// TIA Portal project "GzyHzy_1500" (V15) (continued)
VERSION : 0.1
   VAR
      "1#除尘轴伸端U1相" : Real;   // 临时占位符变量
      "1#除尘轴伸端V1相" : Real;   // 临时占位符变量
      "1#除尘轴伸端W1相" : Real;   // 临时占位符变量
      "1#除尘非轴伸端U2相" : Real;   // 临时占位符变量
      "1#除尘非轴伸端V2相" : Real;   // 临时占位符变量
      "1#除尘非轴伸端W2相" : Real;   // 临时占位符变量
      "1#除尘电机前轴承温度" : Real;   // 临时占位符变量
      "1#除尘电机后轴承温度" : Real;   // 临时占位符变量
      "1#除尘风机前轴承温度" : Real;   // 临时占位符变量
      "1#除尘风机后轴承温度" : Real;   // 临时占位符变量
      DB_VAR10 : Real;   // 临时占位符变量
      DB_VAR11 : Real;   // 临时占位符变量
      DB_VAR12 : Real;   // 临时占位符变量
      DB_VAR13 : Real;   // 临时占位符变量
      DB_VAR14 : Real;   // 临时占位符变量
      DB_VAR15 : Real;   // 临时占位符变量
      DB_VAR16 : Real;   // 临时占位符变量
      DB_VAR17 : Real;   // 临时占位符变量
      DB_VAR18 : Real;   // 临时占位符变量
      DB_VAR19 : Real;   // 临时占位符变量
      DB_VAR20 : Real;   // 临时占位符变量
      DB_VAR21 : Real;   // 临时占位符变量
      DB_VAR22 : Real;   // 临时占位符变量
      DB_VAR23 : Real;   // 临时占位符变量
      DB_VAR24 : Real;   // 临时占位符变量
      DB_VAR25 : Real;   // 临时占位符变量
      DB_VAR26 : Real;   // 临时占位符变量
      DB_VAR27 : Real;   // 临时占位符变量
      DB_VAR28 : Real;   // 临时占位符变量
      DB_VAR29 : Real;   // 临时占位符变量
      DB_VAR30 : Real;   // 临时占位符变量
      DB_VAR31 : Real;   // 临时占位符变量
      DB_VAR32 : Real;   // 临时占位符变量
      DB_VAR33 : Real;   // 临时占位符变量
      DB_VAR34 : Real;   // 临时占位符变量
      DB_VAR35 : Real;   // 临时占位符变量
      DB_VAR36 : Real;   // 临时占位符变量
      DB_VAR37 : Real;   // 临时占位符变量
      DB_VAR38 : Real;   // 临时占位符变量
      DB_VAR39 : Real;   // 临时占位符变量
      DB_VAR40 : Real;   // 临时占位符变量
      DB_VAR41 : Real;   // 临时占位符变量
      DB_VAR42 : Real;   // 临时占位符变量
      DB_VAR43 : Real;   // 临时占位符变量
      DB_VAR44 : Real;   // 临时占位符变量
      DB_VAR45 : Real;   // 临时占位符变量
      DB_VAR46 : Real;   // 临时占位符变量
      DB_VAR47 : Real;   // 临时占位符变量
      DB_VAR48 : Real;   // 临时占位符变量
      DB_VAR49 : Real;   // 临时占位符变量
      "2#除尘轴伸端U1相" : Real;   // 临时占位符变量
      "2#除尘轴伸端V1相" : Real;   // 临时占位符变量
      "2#除尘轴伸端W1相" : Real;   // 临时占位符变量
      "2#除尘非轴伸端U2相" : Real;   // 临时占位符变量
      "2#除尘非轴伸端V2相" : Real;   // 临时占位符变量
      "2#除尘非轴伸端W2相" : Real;   // 临时占位符变量
      "2#除尘电机前轴承温度" : Real;   // 临时占位符变量
      "2#除尘电机后轴承温度" : Real;   // 临时占位符变量
      "2#除尘风机前轴承温度" : Real;   // 临时占位符变量
      "2#除尘风机后轴承温度" : Real;   // 临时占位符变量
      DB_VAR60 : Real;   // 临时占位符变量
      DB_VAR61 : Real;   // 临时占位符变量
      DB_VAR62 : Real;   // 临时占位符变量
      DB_VAR63 : Real;   // 临时占位符变量
      DB_VAR64 : Real;   // 临时占位符变量
      DB_VAR65 : Real;   // 临时占位符变量
      DB_VAR66 : Real;   // 临时占位符变量
   END_VAR
BEGIN
END_DATA_BLOCK

FUNCTION "FC1" : Void   // FC1, LAD
{ S7_Optimized_Access := 'FALSE' }
VERSION : 0.1
BEGIN

REGION Network 1: 1#1号电场二次运行电压
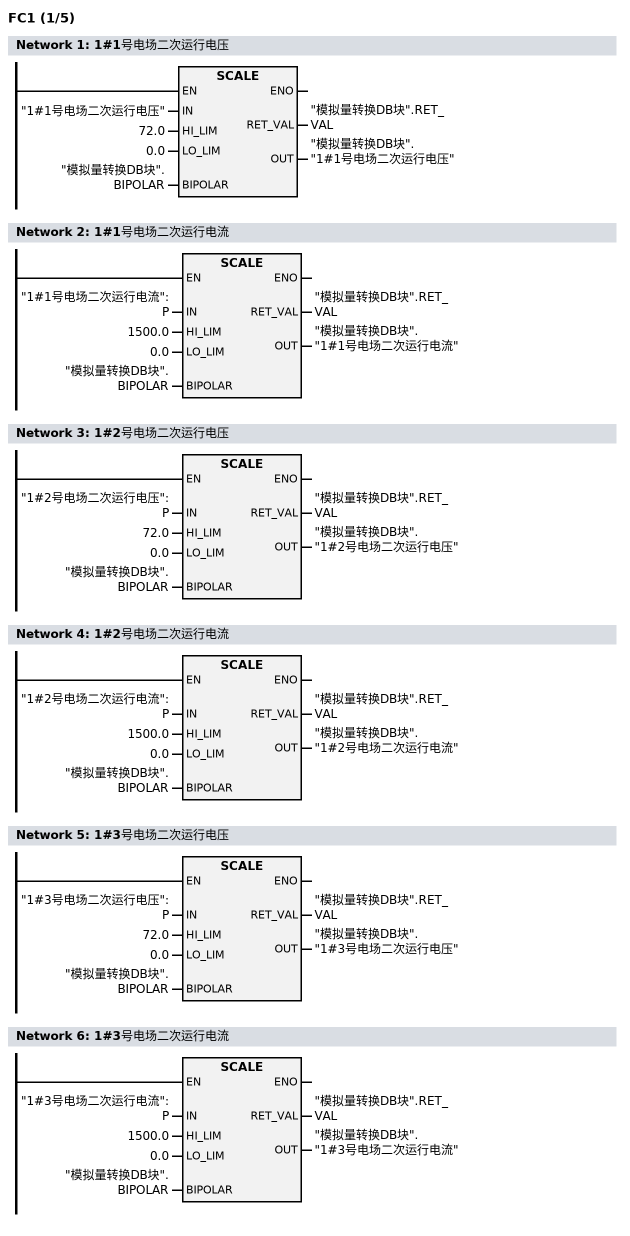
   "模拟量转换DB块".RET_VAL := SCALE(IN := "1#1号电场二次运行电压",
                           HI_LIM := 72.0,
                           LO_LIM := 0.0,
                           BIPOLAR := "模拟量转换DB块".BIPOLAR,
                           OUT => "模拟量转换DB块"."1#1号电场二次运行电压");
END_REGION

REGION Network 2: 1#1号电场二次运行电流
   "模拟量转换DB块".RET_VAL := SCALE(IN := "1#1号电场二次运行电流":P,
                           HI_LIM := 1500.0,
                           LO_LIM := 0.0,
                           BIPOLAR := "模拟量转换DB块".BIPOLAR,
                           OUT => "模拟量转换DB块"."1#1号电场二次运行电流");
END_REGION

REGION Network 3: 1#2号电场二次运行电压
   "模拟量转换DB块".RET_VAL := SCALE(IN := "1#2号电场二次运行电压":P,
                           HI_LIM := 72.0,
                           LO_LIM := 0.0,
                           BIPOLAR := "模拟量转换DB块".BIPOLAR,
                           OUT => "模拟量转换DB块"."1#2号电场二次运行电压");
END_REGION

REGION Network 4: 1#2号电场二次运行电流
   "模拟量转换DB块".RET_VAL := SCALE(IN := "1#2号电场二次运行电流":P,
                           HI_LIM := 1500.0,
                           LO_LIM := 0.0,
                           BIPOLAR := "模拟量转换DB块".BIPOLAR,
                           OUT => "模拟量转换DB块"."1#2号电场二次运行电流");
END_REGION

REGION Network 5: 1#3号电场二次运行电压
   "模拟量转换DB块".RET_VAL := SCALE(IN := "1#3号电场二次运行电压":P,
                           HI_LIM := 72.0,
                           LO_LIM := 0.0,
                           BIPOLAR := "模拟量转换DB块".BIPOLAR,
                           OUT => "模拟量转换DB块"."1#3号电场二次运行电压");
END_REGION

REGION Network 6: 1#3号电场二次运行电流
   "模拟量转换DB块".RET_VAL := SCALE(IN := "1#3号电场二次运行电流":P,
                           HI_LIM := 1500.0,
                           LO_LIM := 0.0,
                           BIPOLAR := "模拟量转换DB块".BIPOLAR,
                           OUT => "模拟量转换DB块"."1#3号电场二次运行电流");
END_REGION

REGION Network 7: 1#4号电场二次运行电压
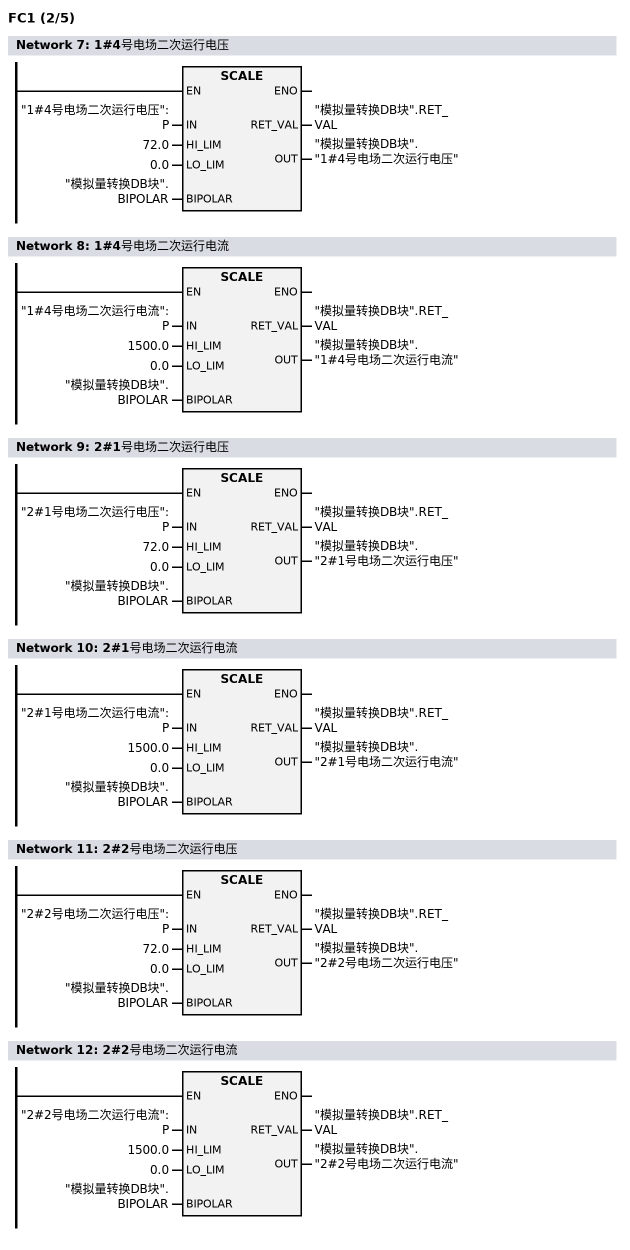
   "模拟量转换DB块".RET_VAL := SCALE(IN := "1#4号电场二次运行电压":P,
                           HI_LIM := 72.0,
                           LO_LIM := 0.0,
                           BIPOLAR := "模拟量转换DB块".BIPOLAR,
                           OUT => "模拟量转换DB块"."1#4号电场二次运行电压");
END_REGION

REGION Network 8: 1#4号电场二次运行电流
   "模拟量转换DB块".RET_VAL := SCALE(IN := "1#4号电场二次运行电流":P,
                           HI_LIM := 1500.0,
                           LO_LIM := 0.0,
                           BIPOLAR := "模拟量转换DB块".BIPOLAR,
                           OUT => "模拟量转换DB块"."1#4号电场二次运行电流");
END_REGION

REGION Network 9: 2#1号电场二次运行电压
   "模拟量转换DB块".RET_VAL := SCALE(IN := "2#1号电场二次运行电压":P,
                           HI_LIM := 72.0,
                           LO_LIM := 0.0,
                           BIPOLAR := "模拟量转换DB块".BIPOLAR,
                           OUT => "模拟量转换DB块"."2#1号电场二次运行电压");
END_REGION

REGION Network 10: 2#1号电场二次运行电流
   "模拟量转换DB块".RET_VAL := SCALE(IN := "2#1号电场二次运行电流":P,
                           HI_LIM := 1500.0,
                           LO_LIM := 0.0,
                           BIPOLAR := "模拟量转换DB块".BIPOLAR,
                           OUT => "模拟量转换DB块"."2#1号电场二次运行电流");
END_REGION

REGION Network 11: 2#2号电场二次运行电压
   "模拟量转换DB块".RET_VAL := SCALE(IN := "2#2号电场二次运行电压":P,
                           HI_LIM := 72.0,
                           LO_LIM := 0.0,
                           BIPOLAR := "模拟量转换DB块".BIPOLAR,
                           OUT => "模拟量转换DB块"."2#2号电场二次运行电压");
END_REGION

REGION Network 12: 2#2号电场二次运行电流
   "模拟量转换DB块".RET_VAL := SCALE(IN := "2#2号电场二次运行电流":P,
                           HI_LIM := 1500.0,
                           LO_LIM := 0.0,
                           BIPOLAR := "模拟量转换DB块".BIPOLAR,
                           OUT => "模拟量转换DB块"."2#2号电场二次运行电流");
END_REGION

REGION Network 13: 2#3号电场二次运行电压
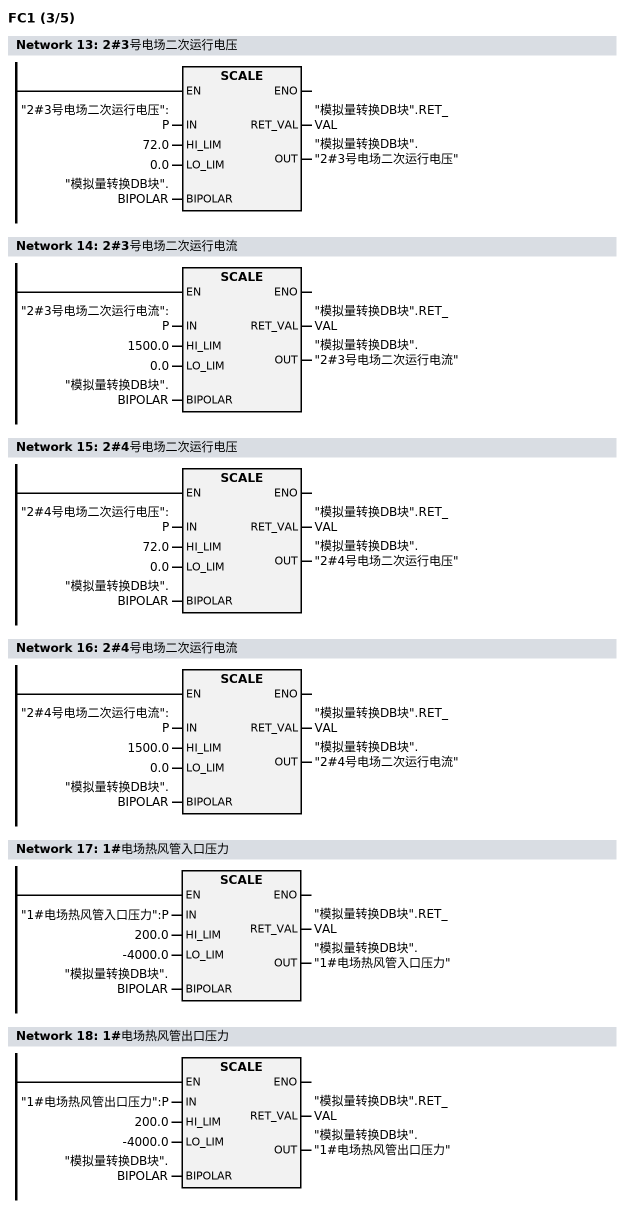
   "模拟量转换DB块".RET_VAL := SCALE(IN := "2#3号电场二次运行电压":P,
                           HI_LIM := 72.0,
                           LO_LIM := 0.0,
                           BIPOLAR := "模拟量转换DB块".BIPOLAR,
                           OUT => "模拟量转换DB块"."2#3号电场二次运行电压");
END_REGION

REGION Network 14: 2#3号电场二次运行电流
   "模拟量转换DB块".RET_VAL := SCALE(IN := "2#3号电场二次运行电流":P,
                           HI_LIM := 1500.0,
                           LO_LIM := 0.0,
                           BIPOLAR := "模拟量转换DB块".BIPOLAR,
                           OUT => "模拟量转换DB块"."2#3号电场二次运行电流");
END_REGION

REGION Network 15: 2#4号电场二次运行电压
   "模拟量转换DB块".RET_VAL := SCALE(IN := "2#4号电场二次运行电压":P,
                           HI_LIM := 72.0,
                           LO_LIM := 0.0,
                           BIPOLAR := "模拟量转换DB块".BIPOLAR,
                           OUT => "模拟量转换DB块"."2#4号电场二次运行电压");
END_REGION

REGION Network 16: 2#4号电场二次运行电流
   "模拟量转换DB块".RET_VAL := SCALE(IN := "2#4号电场二次运行电流":P,
                           HI_LIM := 1500.0,
                           LO_LIM := 0.0,
                           BIPOLAR := "模拟量转换DB块".BIPOLAR,
                           OUT => "模拟量转换DB块"."2#4号电场二次运行电流");
END_REGION

REGION Network 17: 1#电场热风管入口压力
   "模拟量转换DB块".RET_VAL := SCALE(IN := "1#电场热风管入口压力":P,
                           HI_LIM := 200.0,
                           LO_LIM := -4000.0,
                           BIPOLAR := "模拟量转换DB块".BIPOLAR,
                           OUT => "模拟量转换DB块"."1#电场热风管入口压力");
END_REGION

REGION Network 18: 1#电场热风管出口压力
   "模拟量转换DB块".RET_VAL := SCALE(IN := "1#电场热风管出口压力":P,
                           HI_LIM := 200.0,
                           LO_LIM := -4000.0,
                           BIPOLAR := "模拟量转换DB块".BIPOLAR,
                           OUT => "模拟量转换DB块"."1#电场热风管出口压力");
END_REGION

REGION Network 19: 2#电场热风管入口压力
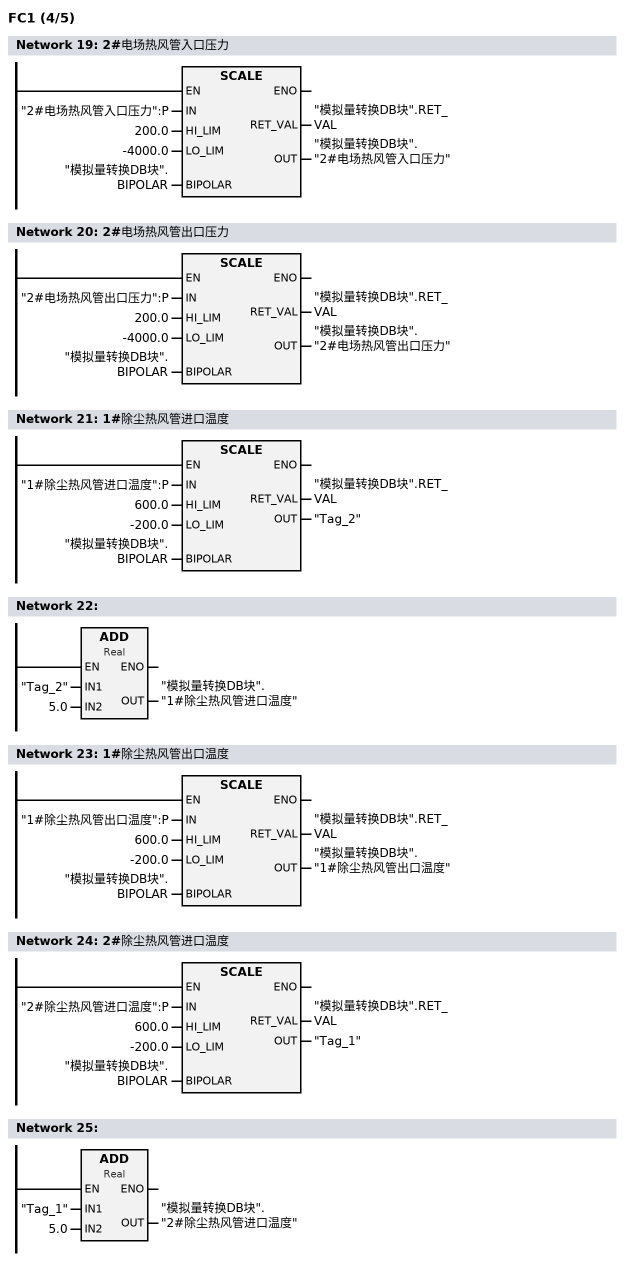
   "模拟量转换DB块".RET_VAL := SCALE(IN := "2#电场热风管入口压力":P,
                           HI_LIM := 200.0,
                           LO_LIM := -4000.0,
                           BIPOLAR := "模拟量转换DB块".BIPOLAR,
                           OUT => "模拟量转换DB块"."2#电场热风管入口压力");
END_REGION

REGION Network 20: 2#电场热风管出口压力
   "模拟量转换DB块".RET_VAL := SCALE(IN := "2#电场热风管出口压力":P,
                           HI_LIM := 200.0,
                           LO_LIM := -4000.0,
                           BIPOLAR := "模拟量转换DB块".BIPOLAR,
                           OUT => "模拟量转换DB块"."2#电场热风管出口压力");
END_REGION

REGION Network 21: 1#除尘热风管进口温度
   "模拟量转换DB块".RET_VAL := SCALE(IN := "1#除尘热风管进口温度":P,
                           HI_LIM := 600.0,
                           LO_LIM := -200.0,
                           BIPOLAR := "模拟量转换DB块".BIPOLAR,
                           OUT => "Tag_2");
END_REGION

REGION Network 22
   RUNG wire#powerrail
      { S7_Templates := "SrcType := Real" } Add(in1 := "Tag_2", in2 := 5.0, out => "模拟量转换DB块"."1#除尘热风管进口温度")
   END_RUNG
   // the same network as SCL:
   "模拟量转换DB块"."1#除尘热风管进口温度" := "Tag_2" + 5.0;
END_REGION

REGION Network 23: 1#除尘热风管出口温度
   "模拟量转换DB块".RET_VAL := SCALE(IN := "1#除尘热风管出口温度":P,
                           HI_LIM := 600.0,
                           LO_LIM := -200.0,
                           BIPOLAR := "模拟量转换DB块".BIPOLAR,
                           OUT => "模拟量转换DB块"."1#除尘热风管出口温度");
END_REGION

REGION Network 24: 2#除尘热风管进口温度
   "模拟量转换DB块".RET_VAL := SCALE(IN := "2#除尘热风管进口温度":P,
                           HI_LIM := 600.0,
                           LO_LIM := -200.0,
                           BIPOLAR := "模拟量转换DB块".BIPOLAR,
                           OUT => "Tag_1");
END_REGION

REGION Network 25
   RUNG wire#powerrail
      { S7_Templates := "SrcType := Real" } Add(in1 := "Tag_1", in2 := 5.0, out => "模拟量转换DB块"."2#除尘热风管进口温度")
   END_RUNG
   // the same network as SCL:
   "模拟量转换DB块"."2#除尘热风管进口温度" := "Tag_1" + 5.0;
END_REGION

REGION Network 26: 2#除尘热风管出口温度
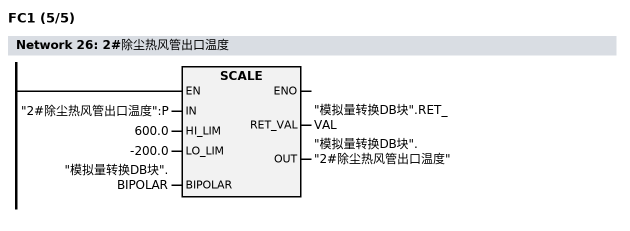
   "模拟量转换DB块".RET_VAL := SCALE(IN := "2#除尘热风管出口温度":P,
                           HI_LIM := 600.0,
                           LO_LIM := -200.0,
                           BIPOLAR := "模拟量转换DB块".BIPOLAR,
                           OUT => "模拟量转换DB块"."2#除尘热风管出口温度");
END_REGION
END_FUNCTION

FUNCTION "DP&MODBUS通讯" : Void   // FC15, LAD
{ S7_Optimized_Access := 'FALSE' }
VERSION : 0.1
BEGIN

REGION Network 1
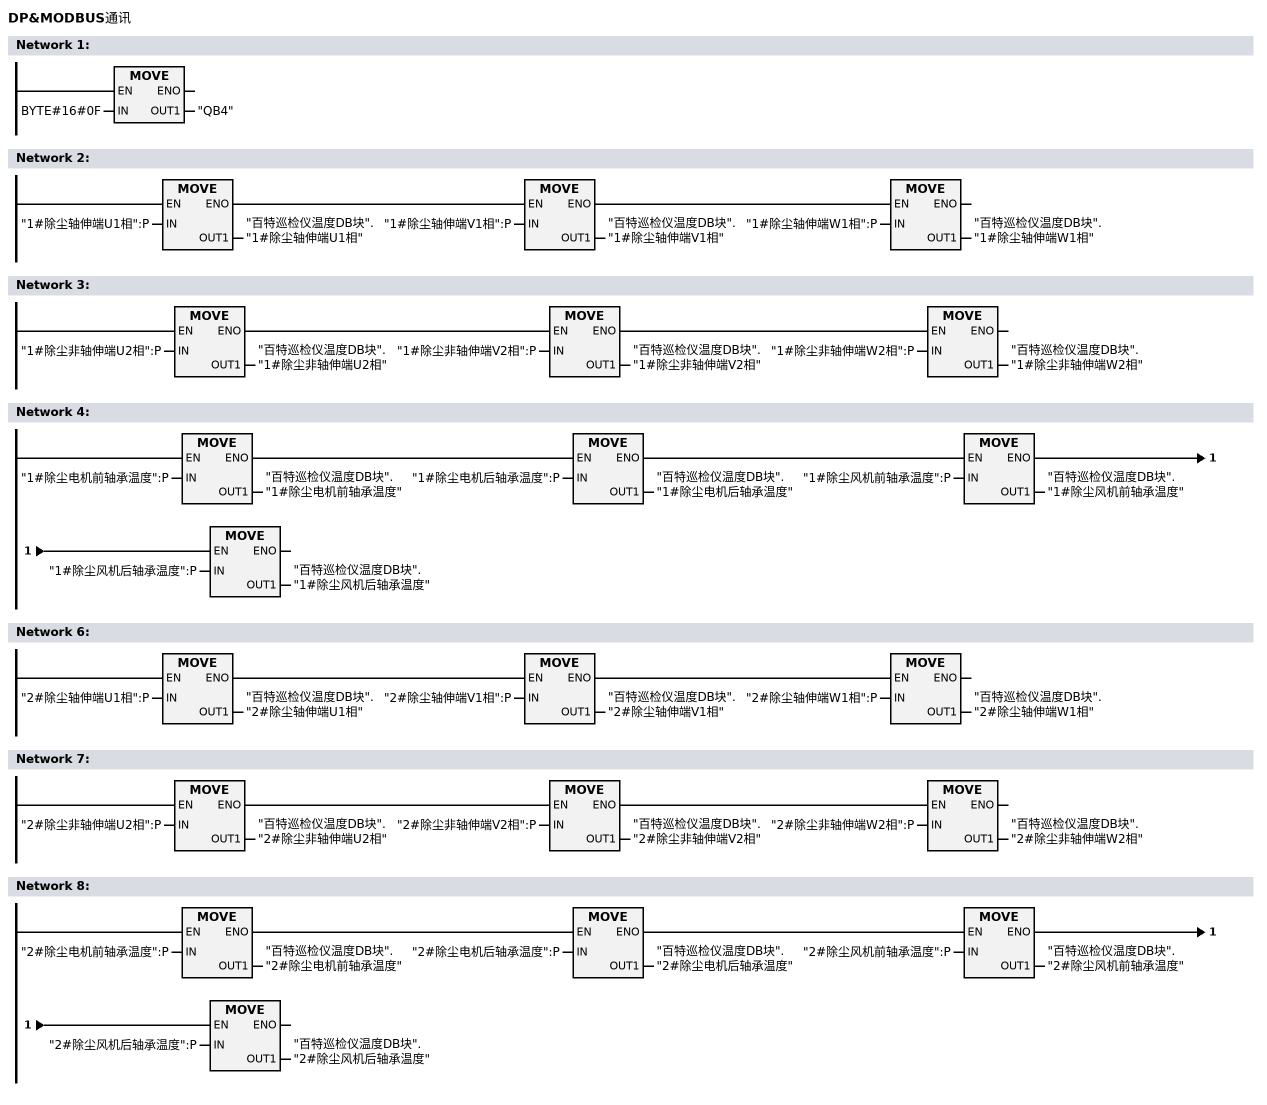
   RUNG wire#powerrail
      { S7_GenerateENO := "TRUE" } Move(in := BYTE#16#0F, out1 => "QB4")
   END_RUNG
   // the same network as SCL:
   "QB4" := BYTE#16#0F;
END_REGION

REGION Network 2
   RUNG wire#powerrail
      { S7_GenerateENO := "TRUE" } Move(in := "1#除尘轴伸端U1相":P, out1 => "百特巡检仪温度DB块"."1#除尘轴伸端U1相")
      { S7_GenerateENO := "TRUE" } Move(in := "1#除尘轴伸端V1相":P, out1 => "百特巡检仪温度DB块"."1#除尘轴伸端V1相")
      { S7_GenerateENO := "TRUE" } Move(in := "1#除尘轴伸端W1相":P, out1 => "百特巡检仪温度DB块"."1#除尘轴伸端W1相")
   END_RUNG
   // the same network as SCL:
   // ENO of a box is taken as its EN; it also drops when the box reports an error
   "百特巡检仪温度DB块"."1#除尘轴伸端U1相" := "1#除尘轴伸端U1相":P;
   "百特巡检仪温度DB块"."1#除尘轴伸端V1相" := "1#除尘轴伸端V1相":P;
   "百特巡检仪温度DB块"."1#除尘轴伸端W1相" := "1#除尘轴伸端W1相":P;
END_REGION

REGION Network 3
   RUNG wire#powerrail
      { S7_GenerateENO := "TRUE" } Move(in := "1#除尘非轴伸端U2相":P, out1 => "百特巡检仪温度DB块"."1#除尘非轴伸端U2相")
      { S7_GenerateENO := "TRUE" } Move(in := "1#除尘非轴伸端V2相":P, out1 => "百特巡检仪温度DB块"."1#除尘非轴伸端V2相")
      { S7_GenerateENO := "TRUE" } Move(in := "1#除尘非轴伸端W2相":P, out1 => "百特巡检仪温度DB块"."1#除尘非轴伸端W2相")
   END_RUNG
   // the same network as SCL:
   // ENO of a box is taken as its EN; it also drops when the box reports an error
   "百特巡检仪温度DB块"."1#除尘非轴伸端U2相" := "1#除尘非轴伸端U2相":P;
   "百特巡检仪温度DB块"."1#除尘非轴伸端V2相" := "1#除尘非轴伸端V2相":P;
   "百特巡检仪温度DB块"."1#除尘非轴伸端W2相" := "1#除尘非轴伸端W2相":P;
END_REGION

REGION Network 4
   RUNG wire#powerrail
      { S7_GenerateENO := "TRUE" } Move(in := "1#除尘电机前轴承温度":P, out1 => "百特巡检仪温度DB块"."1#除尘电机前轴承温度")
      { S7_GenerateENO := "TRUE" } Move(in := "1#除尘电机后轴承温度":P, out1 => "百特巡检仪温度DB块"."1#除尘电机后轴承温度")
      { S7_GenerateENO := "TRUE" } Move(in := "1#除尘风机前轴承温度":P, out1 => "百特巡检仪温度DB块"."1#除尘风机前轴承温度")
      { S7_GenerateENO := "TRUE" } Move(in := "1#除尘风机后轴承温度":P, out1 => "百特巡检仪温度DB块"."1#除尘风机后轴承温度")
   END_RUNG
   // the same network as SCL:
   // ENO of a box is taken as its EN; it also drops when the box reports an error
   "百特巡检仪温度DB块"."1#除尘电机前轴承温度" := "1#除尘电机前轴承温度":P;
   "百特巡检仪温度DB块"."1#除尘电机后轴承温度" := "1#除尘电机后轴承温度":P;
   "百特巡检仪温度DB块"."1#除尘风机前轴承温度" := "1#除尘风机前轴承温度":P;
   "百特巡检仪温度DB块"."1#除尘风机后轴承温度" := "1#除尘风机后轴承温度":P;
END_REGION

REGION Network 6
   RUNG wire#powerrail
      { S7_GenerateENO := "TRUE" } Move(in := "2#除尘轴伸端U1相":P, out1 => "百特巡检仪温度DB块"."2#除尘轴伸端U1相")
      { S7_GenerateENO := "TRUE" } Move(in := "2#除尘轴伸端V1相":P, out1 => "百特巡检仪温度DB块"."2#除尘轴伸端V1相")
      { S7_GenerateENO := "TRUE" } Move(in := "2#除尘轴伸端W1相":P, out1 => "百特巡检仪温度DB块"."2#除尘轴伸端W1相")
   END_RUNG
   // the same network as SCL:
   // ENO of a box is taken as its EN; it also drops when the box reports an error
   "百特巡检仪温度DB块"."2#除尘轴伸端U1相" := "2#除尘轴伸端U1相":P;
   "百特巡检仪温度DB块"."2#除尘轴伸端V1相" := "2#除尘轴伸端V1相":P;
   "百特巡检仪温度DB块"."2#除尘轴伸端W1相" := "2#除尘轴伸端W1相":P;
END_REGION

REGION Network 7
   RUNG wire#powerrail
      { S7_GenerateENO := "TRUE" } Move(in := "2#除尘非轴伸端U2相":P, out1 => "百特巡检仪温度DB块"."2#除尘非轴伸端U2相")
      { S7_GenerateENO := "TRUE" } Move(in := "2#除尘非轴伸端V2相":P, out1 => "百特巡检仪温度DB块"."2#除尘非轴伸端V2相")
      { S7_GenerateENO := "TRUE" } Move(in := "2#除尘非轴伸端W2相":P, out1 => "百特巡检仪温度DB块"."2#除尘非轴伸端W2相")
   END_RUNG
   // the same network as SCL:
   // ENO of a box is taken as its EN; it also drops when the box reports an error
   "百特巡检仪温度DB块"."2#除尘非轴伸端U2相" := "2#除尘非轴伸端U2相":P;
   "百特巡检仪温度DB块"."2#除尘非轴伸端V2相" := "2#除尘非轴伸端V2相":P;
   "百特巡检仪温度DB块"."2#除尘非轴伸端W2相" := "2#除尘非轴伸端W2相":P;
END_REGION

REGION Network 8
   RUNG wire#powerrail
      { S7_GenerateENO := "TRUE" } Move(in := "2#除尘电机前轴承温度":P, out1 => "百特巡检仪温度DB块"."2#除尘电机前轴承温度")
      { S7_GenerateENO := "TRUE" } Move(in := "2#除尘电机后轴承温度":P, out1 => "百特巡检仪温度DB块"."2#除尘电机后轴承温度")
      { S7_GenerateENO := "TRUE" } Move(in := "2#除尘风机前轴承温度":P, out1 => "百特巡检仪温度DB块"."2#除尘风机前轴承温度")
      { S7_GenerateENO := "TRUE" } Move(in := "2#除尘风机后轴承温度":P, out1 => "百特巡检仪温度DB块"."2#除尘风机后轴承温度")
   END_RUNG
   // the same network as SCL:
   // ENO of a box is taken as its EN; it also drops when the box reports an error
   "百特巡检仪温度DB块"."2#除尘电机前轴承温度" := "2#除尘电机前轴承温度":P;
   "百特巡检仪温度DB块"."2#除尘电机后轴承温度" := "2#除尘电机后轴承温度":P;
   "百特巡检仪温度DB块"."2#除尘风机前轴承温度" := "2#除尘风机前轴承温度":P;
   "百特巡检仪温度DB块"."2#除尘风机后轴承温度" := "2#除尘风机后轴承温度":P;
END_REGION
END_FUNCTION

ORGANIZATION_BLOCK "Main"   // OB1, LAD, ProgramCycle
TITLE = "Main Program Sweep (Cycle)"
{ S7_Optimized_Access := 'TRUE' }
VERSION : 0.1
   VAR_INPUT
      Initial_Call : Bool;   // Initial call of this OB
      Remanence : Bool;   // =True, if remanent data are available
   END_VAR
BEGIN

REGION Network 1
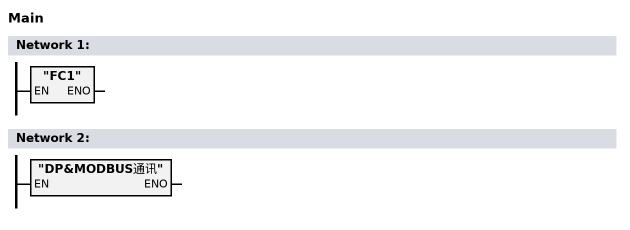
   RUNG wire#powerrail
      "FC1"()
   END_RUNG
   // the same network as SCL:
   "FC1"();
END_REGION

REGION Network 2
   RUNG wire#powerrail
      "DP&MODBUS通讯"()
   END_RUNG
   // the same network as SCL:
   "DP&MODBUS通讯"();
END_REGION
END_ORGANIZATION_BLOCK

// ===== PLC "1#GZY"  CPU 1511-1 PN =====

VAR_GLOBAL   // PLC tag table "默认变量表"
   "1#干燥窑主机远程" AT %I0.0 : Bool;
   "1#干燥窑主机变频备妥" AT %I0.1 : Bool;
   "1#干燥窑主机散热风机运行" AT %I0.2 : Bool;
   "1#干燥窑变频运行" AT %I0.3 : Bool;
   "1#干燥窑变频故障" AT %I0.4 : Bool;
   "1#干燥窑稀油中控" AT %I1.0 : Bool;
   "1#干燥窑稀油1#泵运行" AT %I1.1 : Bool;
   "1#干燥窑稀油2#泵运行" AT %I1.2 : Bool;
   "1#干燥窑稀油油差下限" AT %I1.3 : Bool;
   "1#干燥窑稀油油位上限" AT %I1.4 : Bool;
   "1#干燥窑稀油油位下限" AT %I1.5 : Bool;
   "1#干燥窑稀油1#泵故障" AT %I1.6 : Bool;
   "1#干燥窑稀油2#泵故障" AT %I1.7 : Bool;
   "1#干燥窑挡轮备妥" AT %I2.0 : Bool;
   "1#干燥窑挡轮1#泵运行" AT %I2.1 : Bool;
   "1#干燥窑挡轮2#泵运行" AT %I2.2 : Bool;
   "1#干燥窑挡轮溢流阀运行" AT %I2.3 : Bool;
   "1#干燥窑挡轮行程过低" AT %I2.4 : Bool;
   "1#干燥窑挡轮故障" AT %I2.5 : Bool;
   "1#皮带_湿矿上料皮带中控" AT %I3.0 : Bool;
   "1#皮带_湿矿上料皮带运行" AT %I3.1 : Bool;
   "1#皮带_湿矿上料皮带故障" AT %I3.2 : Bool;
   "2#皮带_湿矿转1#干燥窑皮带中控" AT %I3.3 : Bool;
   "2#皮带_湿矿转1#干燥窑皮带运行" AT %I3.4 : Bool;
   "2#皮带_湿矿转1#干燥窑皮带故障" AT %I3.5 : Bool;
   "4#皮带_干矿下料皮带中控" AT %I4.0 : Bool;
   "4#皮带_干矿下料皮带运行" AT %I4.1 : Bool;
   "4#皮带_干矿下料皮带故障" AT %I4.2 : Bool;
   "5#皮带_干矿下料转破碎皮带中控" AT %I4.3 : Bool;
   "5#皮带_干矿下料转破碎皮带运行" AT %I4.4 : Bool;
   "5#皮带_干矿下料转破碎皮带故障" AT %I4.5 : Bool;
   "6#皮带_破碎提升中转皮带中控" AT %I5.0 : Bool;
   "6#皮带_破碎提升中转皮带运行" AT %I5.1 : Bool;
   "6#皮带_破碎提升中转皮带故障" AT %I5.2 : Bool;
   "7#皮带_中转到干矿棚皮带中控" AT %I5.3 : Bool;
   "7#皮带_中转到干矿棚皮带运行" AT %I5.4 : Bool;
   "7#皮带_中转到干矿棚皮带故障" AT %I5.5 : Bool;
   "定量给煤机中控" AT %I6.3 : Bool;
   "定量给煤机运行" AT %I6.4 : Bool;
   "定量给煤机故障" AT %I6.5 : Bool;
   "定量给煤机流量脉冲" AT %I6.6 : Bool;
   "煤粉仓收尘风机中控" AT %I7.0 : Bool;
   "煤粉仓收尘风机运行" AT %I7.1 : Bool;
   "煤粉仓收尘风机故障" AT %I7.2 : Bool;
   "1#干燥窑一次风机中控" AT %I8.0 : Bool;
   "1#干燥窑一次风机运行" AT %I8.1 : Bool;
   "1#干燥窑一次风机故障" AT %I8.2 : Bool;
   "1#干燥窑二次风机中控" AT %I8.3 : Bool;
   "1#干燥窑二次风机运行" AT %I8.4 : Bool;
   "1#干燥窑二次风机故障" AT %I8.5 : Bool;
   "1#干燥窑备用一次风机中控" AT %I9.0 : Bool;
   "1#干燥窑备用一次风机运行" AT %I9.1 : Bool;
   "1#干燥窑备用一次风机故障" AT %I9.2 : Bool;
   "1#干燥窑备用二次风机中控" AT %I9.3 : Bool;
   "1#干燥窑备用二次风机运行" AT %I9.4 : Bool;
   "1#干燥窑备用二次风机故障" AT %I9.5 : Bool;
   "1#干燥窑振动筛中控" AT %I10.0 : Bool;
   "1#干燥窑振动筛运行" AT %I10.1 : Bool;
   "1#干燥窑振动筛故障" AT %I10.2 : Bool;
   "1#干燥窑破碎机中控" AT %I10.4 : Bool;
   "1#干燥窑破碎机运行" AT %I10.5 : Bool;
   "1#干燥窑破碎机故障" AT %I10.6 : Bool;
   "1#干燥窑主传动转速" AT %IW256 : Int;
   "1#干燥窑主传动电流" AT %IW258 : Int;
   "1#干燥窑二次风机电流" AT %IW260 : Int;
   "1#干燥窑一次风机电流" AT %IW262 : Int;
   "1#干燥窑二次风机频率" AT %IW264 : Int;
   "1#干燥窑窑尾压力" AT %IW266 : Int;
   "1#干燥窑备用一次风机频率" AT %IW268 : Int;
   "1#干燥窑备用一次风机电流" AT %IW270 : Int;
   "1#干燥窑备用二次风机频率" AT %IW272 : Int;
   "1#干燥窑备用二次风机电流" AT %IW274 : Int;
   "定量给煤机流量" AT %IW276 : Int;
   "烟气管道进口压力" AT %IW278 : Int;
   "1#干燥窑一次风压" AT %IW280 : Int;
   "1#干燥窑二次风压" AT %IW282 : Int;
   "煤粉仓压力" AT %IW284 : Int;
   "混合室压力" AT %IW286 : Int;
   "煤粉仓温度1(PT100)" AT %IW288 : Int;
   "煤粉仓温度2(PT100)" AT %IW290 : Int;
   "煤粉仓温度3(PT100)" AT %IW292 : Int;
   "煤粉仓温度4(PT100)" AT %IW294 : Int;
   "窑尾温度 K偶" AT %IW296 : Int;
   "烟气管道进口温度 K偶" AT %IW298 : Int;
   "燃烧室温度 4~20mA" AT %IW300 : Int;
   "混合室温度 4~20mA" AT %IW302 : Int;
   "1#干燥窑断路器合闸" AT %I0.5 : Bool;
   "1#干燥窑断路器分闸" AT %I0.6 : Bool;
   "1#干燥窑进料口压力" AT %IW304 : Int;
   "1#窑主电机B相绕组温度" AT %ID388 : Real;
   "1#窑主电机C相绕组温度" AT %ID392 : Real;
   "1#窑主电机前轴承温度" AT %ID396 : Real;
   "1#窑主电机后轴承温度" AT %ID400 : Real;
   "I0_7" AT %I0.7 : Bool;
   "I2_6" AT %I2.6 : Bool;
   "I2_7" AT %I2.7 : Bool;
   "I3_6" AT %I3.6 : Bool;
   "I3_7" AT %I3.7 : Bool;
   "I4_6" AT %I4.6 : Bool;
   "I4_7" AT %I4.7 : Bool;
   "I5_6" AT %I5.6 : Bool;
   "I5_7" AT %I5.7 : Bool;
   "I6_0" AT %I6.0 : Bool;
   "I6_1" AT %I6.1 : Bool;
   "I6_2" AT %I6.2 : Bool;
   "I6_7" AT %I6.7 : Bool;
   "I7_3" AT %I7.3 : Bool;
   "I7_4" AT %I7.4 : Bool;
   "I7_5" AT %I7.5 : Bool;
   "I7_6" AT %I7.6 : Bool;
   "I7_7" AT %I7.7 : Bool;
   "I8_6" AT %I8.6 : Bool;
   "I8_7" AT %I8.7 : Bool;
   "I9_6" AT %I9.6 : Bool;
   "I9_7" AT %I9.7 : Bool;
   "I10_3" AT %I10.3 : Bool;
   "I10_7" AT %I10.7 : Bool;
   "8#皮带_中转到干矿棚皮带2中控" AT %I11.0 : Bool;
   "8#皮带_中转到干矿棚皮带2运行" AT %I11.1 : Bool;
   "8#皮带_中转到干矿棚皮带2故障" AT %I11.2 : Bool;
   "I11_3" AT %I11.3 : Bool;
   "I11_4" AT %I11.4 : Bool;
   "I11_5" AT %I11.5 : Bool;
   "I11_6" AT %I11.6 : Bool;
   "I11_7" AT %I11.7 : Bool;
   "1#给煤机出料口负压" AT %IW306 : Int;
   "振动筛转速" AT %IW308 : Int;
   "振动筛电流" AT %IW310 : Int;
   "PIW312" AT %IW312 : Int;
   "PIW314" AT %IW314 : Int;
   "PIW316" AT %IW316 : Int;
   "PIW318" AT %IW318 : Int;
   "1#窑A档轴温1" AT %ID320 : Real;
   "1#窑A档油温1" AT %ID324 : Real;
   "1#窑A档轴温2" AT %ID328 : Real;
   "1#窑A档油温2" AT %ID332 : Real;
   "1#窑A档轴温3" AT %ID336 : Real;
   "1#窑A档油温3" AT %ID340 : Real;
   "1#窑A档轴温4" AT %ID344 : Real;
   "1#窑A档油温4" AT %ID348 : Real;
   "1#窑B档轴温1" AT %ID352 : Real;
   "1#窑B档油温1" AT %ID356 : Real;
   "1#窑B档轴温2" AT %ID360 : Real;
   "1#窑B档油温2" AT %ID364 : Real;
   "1#窑B档轴温3" AT %ID368 : Real;
   "1#窑B档油温3" AT %ID372 : Real;
   "1#窑B档轴温4" AT %ID376 : Real;
   "1#窑B档油温4" AT %ID380 : Real;
   "1#窑主电机A相绕组温度" AT %ID384 : Real;
   "1#干燥窑煤粉仓称重" AT %ID440 : Real;
   "Tag_11" AT %ID412 : DWord;
   "干燥窑主机风机合闸" AT %Q0.0 : Bool;
   "干燥窑主传动分闸" AT %Q0.1 : Bool;
   "干燥窑主传动变频启动" AT %Q0.2 : Bool;
   "干燥窑主传稀油站启动" AT %Q0.3 : Bool;
   "湿矿上料皮带启动  (1#皮带)" AT %Q0.4 : Bool;
   "湿矿转1#干燥窑皮带启动  (2#皮带)" AT %Q0.5 : Bool;
   "干矿下料皮带启动  (4#皮带)" AT %Q0.6 : Bool;
   "干矿下料转破碎皮带启动  (5#皮带)" AT %Q0.7 : Bool;
   "破碎提升中转皮带启动  (6#皮带)" AT %Q1.0 : Bool;
   "定量给煤机启动" AT %Q1.2 : Bool;
   "煤粉仓收尘风机启动" AT %Q1.3 : Bool;
   "干矿破碎启动" AT %Q1.4 : Bool;
   "振动筛启动" AT %Q1.5 : Bool;
   "干燥窑挡轮油站启动" AT %Q1.6 : Bool;
   "1#干燥窑一次风机启动" AT %Q2.0 : Bool;
   "1#干燥窑二次风机启动" AT %Q2.1 : Bool;
   "1#干燥窑备用一次风机启动" AT %Q2.2 : Bool;
   "1#干燥窑备用二次风机启动" AT %Q2.3 : Bool;
   "Tag_8" AT %QB4 : Byte;
   "1#干燥窑转速给定" AT %QW256 : Int;
   "定量给煤机流量给定" AT %QW258 : Int;
   "PQW264" AT %QW264 : Int;
   "1#干燥窑二次风机频率给定" AT %QW266 : Int;
   "PQW268" AT %QW268 : Int;
   "1#干燥窑备用二次风机频率给定" AT %QW270 : Int;
   "中转到干矿棚皮带启动  (7#皮带)" AT %Q1.1 : Bool;
   "中转到干矿棚皮带2启动  (8#皮带)" AT %Q1.7 : Bool;
   "Q2_4" AT %Q2.4 : Bool;
   "Q2_5" AT %Q2.5 : Bool;
   "Q2_6" AT %Q2.6 : Bool;
   "Q2_7" AT %Q2.7 : Bool;
   "Q3_0" AT %Q3.0 : Bool;
   "Q3_1" AT %Q3.1 : Bool;
   "Q3_2" AT %Q3.2 : Bool;
   "Q3_3" AT %Q3.3 : Bool;
   "Q3_4" AT %Q3.4 : Bool;
   "Q3_5" AT %Q3.5 : Bool;
   "Q3_6" AT %Q3.6 : Bool;
   "Q3_7" AT %Q3.7 : Bool;
   "振动筛转速给定" AT %QW260 : Int;
   "Tag_1" AT %MW4 : Word;
   "Tag_2" AT %M400.0 : Bool;
   "连锁解锁" AT %M400.2 : Bool;
   "干燥窑连锁信号" AT %M400.3 : Bool;
   "Tag_4" AT %M400.5 : Bool;
   "Tag_5" AT %MW410 : Word;
   "Tag_6" AT %MW412 : Word;
   "Tag_32" AT %M1001.0 : Bool;
   "Clock_Byte" AT %MB0 : Byte;
   "Clock_10Hz" AT %M0.0 : Bool;
   "Clock_5Hz" AT %M0.1 : Bool;
   "Clock_2.5Hz" AT %M0.2 : Bool;
   "Clock_2Hz" AT %M0.3 : Bool;
   "Clock_1.25Hz" AT %M0.4 : Bool;
   "Clock_1Hz" AT %M0.5 : Bool;
   "Clock_0.625Hz" AT %M0.6 : Bool;
   "Clock_0.5Hz" AT %M0.7 : Bool;
   "System_Byte" AT %MB1 : Byte;
   "FirstScan" AT %M1.0 : Bool;
   "DiagStatusUpdate" AT %M1.1 : Bool;
   "AlwaysTRUE" AT %M1.2 : Bool;
   "AlwaysFALSE" AT %M1.3 : Bool;
   "Tag_9" AT %M99.0 : Bool;
   "8#皮带_中转到干矿棚皮带2画面启动" AT %M10.0 : Bool;
   "8#皮带_中转到干矿棚皮带2画面停止" AT %M10.1 : Bool;
   "Tag_12" AT %M500.0 : Bool;
   "稀油站油压长时间低" AT %T6 : Timer;
   "稀油站启动10S" AT %T7 : Timer;
   "稀油站油差下限时间" AT %T8 : Timer;
   "Tag_41" AT %T1 : Timer;
   "Tag_42" AT %T2 : Timer;
   "干燥窑稀油站故障延时" AT %T3 : Timer;
   "Tag_10" AT %T10 : Timer;
   "Tag_3" AT %C1 : Counter;
   "Tag_7" AT %C2 : Counter;
END_VAR

DATA_BLOCK "驱动"   // DB1
{ S7_Optimized_Access := 'FALSE' }
VERSION : 0.1
   VAR
      "1#二次风机启动" : Bool;
      "1#二次风机停止" : Bool;
      "1#干燥窑主机合闸" : Bool;
      "1#干燥窑主机分闸" : Bool;
      "1#备用二次风机启动" : Bool;
      "1#备用二次风机停止" : Bool;
      "1#干燥窑主机启动" : Bool;
      "1#干燥窑主机停止" : Bool;
      "gzy1#湿矿皮带启动1#皮带" : Bool;
      "gzy1#湿矿皮带停止1#皮带" : Bool;
      "gzy进窑1#皮带启动2#皮带" : Bool;
      "gzy进窑1#皮带启动2#皮带_1" : Bool;
      STAT12 : Bool;
      STAT13 : Bool;
      "gzy干矿下料皮带启动4#皮带" : Bool;
      "gzy干矿下料皮带启动4#皮带_1" : Bool;
      "gzy干矿提升到破碎启动5#皮带" : Bool;
      "gzy干矿提升到破碎停止5#皮带" : Bool;
      破碎机启动 : Bool;
      破碎机停止 : Bool;
      振动筛启动 : Bool;
      振动筛停止 : Bool;
      "破碎到中转皮带启动6#皮带" : Bool;
      "破碎到中转皮带停止6#皮带" : Bool;
      "中转干矿棚皮带启动7#皮带" : Bool;
      "中转干矿棚皮带停止7#皮带" : Bool;
      STAT26 : Bool;
      STAT27 : Bool;
      "1#一次风机启动" : Bool;
      "1#一次风机停止" : Bool;
      "1#备用一次风机启动" : Bool;
      "1#备用一次风机停止" : Bool;
      STAT32 : Bool;
      STAT33 : Bool;
      "1#干燥窑煤粉收尘风机启动" : Bool;
      "1#干燥窑煤粉收尘风机停止" : Bool;
      "1#干燥窑锁风给煤机启动" : Bool;
      "1#干燥窑锁风给煤机停止" : Bool;
      "1#干燥窑给煤机分割轮启动" : Bool;
      "1#干燥窑给煤机分割轮停止" : Bool;
      STAT40 : Bool;
      STAT41 : Bool;
      STAT42 : Bool;
      STAT43 : Bool;
      STAT44 : Bool;
      STAT45 : Bool;
      STAT46 : Bool;
      STAT47 : Bool;
      STAT48 : Bool;
      STAT49 : Bool;
      STAT50 : Bool;
      STAT51 : Bool;
      STAT52 : Bool;
      STAT53 : Bool;
      STAT54 : Bool;
      STAT55 : Bool;
      STAT56 : Bool;
      "1#干燥窑联锁解锁" : Bool;
      "1#干燥窑定量给煤机班累计清零" : Bool;
      "1#干燥窑定量给煤机日累计清零" : Bool;
      "1#干燥窑定量给煤机总累计清零" : Bool;
      STAT61 : Bool;
      STAT62 : Bool;
      STAT63 : Bool;
      "1#干燥窑稀油站启动" : Bool;
      "1#干燥窑稀油站停止" : Bool;
      STAT66 : Bool;
      STAT67 : Bool;
      "1#干燥窑挡轮油站启动" : Bool;
      "1#干燥窑挡轮油站停止" : Bool;
      STAT68 : Bool;
      STAT69 : Bool;
   END_VAR
BEGIN
END_DATA_BLOCK
